HMI tags "Default tag table"
   "10_DI_DATA_5T1_PWR_OK" : Bool = PLC "10_DI_DATA".5T1_PWR_OK, 1 s
   "10_DI_DATA_6Q6_PWR_OK" : Bool = PLC "10_DI_DATA".6Q6_PWR_OK, 1 s
   "10_DI_DATA_CV341_CLSD" : Bool = PLC "10_DI_DATA".CV341_CLSD, 1 s
   "10_DI_DATA_CV341_OPN" : Bool = PLC "10_DI_DATA".CV341_OPN, 1 s
   "10_DI_DATA_CV358_CLSD" : Bool = PLC "10_DI_DATA".CV358_CLSD, 1 s
   "10_DI_DATA_CV358_OPN" : Bool = PLC "10_DI_DATA".CV358_OPN, 1 s
   "10_DI_DATA_CV406_CLSD" : Bool = PLC "10_DI_DATA".CV406_CLSD, 1 s
   "10_DI_DATA_CV406_OPN" : Bool = PLC "10_DI_DATA".CV406_OPN, 1 s
   "10_DI_DATA_CV407_CLSD" : Bool = PLC "10_DI_DATA".CV407_CLSD, 1 s
   "10_DI_DATA_CV407_OPN" : Bool = PLC "10_DI_DATA".CV407_OPN, 1 s
   "10_DI_DATA_CV409_CLSD" : Bool = PLC "10_DI_DATA".CV409_CLSD, 1 s
   "10_DI_DATA_CV409_OPN" : Bool = PLC "10_DI_DATA".CV409_OPN, 1 s
   "10_DI_DATA_CV411_CLSD" : Bool = PLC "10_DI_DATA".CV411_CLSD, 1 s
   "10_DI_DATA_CV411_OPN" : Bool = PLC "10_DI_DATA".CV411_OPN, 1 s
   "10_DI_DATA_CV441_CLSD" : Bool = PLC "10_DI_DATA".CV441_CLSD, 1 s
   "10_DI_DATA_CV441_OPN" : Bool = PLC "10_DI_DATA".CV441_OPN, 1 s
   "10_DI_DATA_E_400_NOK" : Bool = PLC "10_DI_DATA".E_400_NOK, 1 s
   "10_DI_DATA_E_400_RUN" : Bool = PLC "10_DI_DATA".E_400_RUN, 1 s
   "10_DI_DATA_E_400_SHTDN" : Bool = PLC "10_DI_DATA".E_400_SHTDN, 1 s
   "10_DI_DATA_E_400_STPD" : Bool = PLC "10_DI_DATA".E_400_STPD, 1 s
   "10_DI_DATA_EPB_8S1" : Bool = PLC "10_DI_DATA".EPB_8S1, 1 s
   "10_DI_DATA_FS_332 FLW_OK" : Bool = PLC "10_DI_DATA"."FS_332 FLW_OK", 1 s
   "10_DI_DATA_FS_350_FLW_OK" : Bool = PLC "10_DI_DATA".FS_350_FLW_OK, 1 s
   "10_DI_DATA_LS_303_LO" : Bool = PLC "10_DI_DATA".LS_303_LO, 1 s
   "10_DI_DATA_P_303_ENBLD" : Bool = PLC "10_DI_DATA".P_303_ENBLD, 1 s
   "10_DI_DATA_P_303_OK" : Bool = PLC "10_DI_DATA".P_303_OK, 1 s
   "10_DI_DATA_P_304_ENBLD" : Bool = PLC "10_DI_DATA".P_304_ENBLD, 1 s
   "10_DI_DATA_P_304_OK" : Bool = PLC "10_DI_DATA".P_304_OK, 1 s
   "10_DI_DATA_PB_10S1" : Bool = PLC "10_DI_DATA".PB_10S1, 1 s
   "10_DI_DATA_PB_10S2" : Bool = PLC "10_DI_DATA".PB_10S2, 1 s
   "10_DI_DATA_R3_SPR_DI_136_0" : Bool = PLC "10_DI_DATA".R3_SPR_DI_136_0, 1 s
   "10_DI_DATA_R3_SPR_DI_136_1" : Bool = PLC "10_DI_DATA".R3_SPR_DI_136_1, 1 s
   "100_BC_AUTO_SEQ_DB_CRNT_STEP" : Int = PLC "100_BC_AUTO_SEQ_DB".CRNT_STEP, 1 s
   "100_GCU_AUTO_SEQ_DB_CRNT_STEP" : Int = PLC "100_GCU_AUTO_SEQ_DB".CRNT_STEP, 1 s
   "100_GCU_AUTO_SEQ_DB_RNG" : Bool = PLC "100_GCU_AUTO_SEQ_DB".RNG, 1 s
   "100_IGG_AUTO_SEQ_DB_CRNT_STEP" : Int = PLC "100_IGG_AUTO_SEQ_DB".CRNT_STEP, 1 s
   "101_Fuel_Pumps_DB_Duty Is A" : Bool = PLC "101_Fuel_Pumps_DB"."Duty Is A", 1 s
   "101_Fuel_Pumps_DB_Duty Is B" : Bool = PLC "101_Fuel_Pumps_DB"."Duty Is B", 1 s
   "102_Pilot_Burner_DB_RUNNING" : Bool = PLC "102_Pilot_Burner_DB".RUNNING, 1 s
   "103_Main_Burner_DB_Days burn_CV" : Int = PLC "103_Main_Burner_DB"."Days burn".CV, 1 s
   "103_Main_Burner_DB_DN_OK" : Bool = PLC "103_Main_Burner_DB".DN_OK, 1 s
   "103_Main_Burner_DB_Hours burn_CV" : Int = PLC "103_Main_Burner_DB"."Hours burn".CV, 1 s
   "103_Main_Burner_DB_Minutes burn_CV" : Int = PLC "103_Main_Burner_DB"."Minutes burn".CV, 1 s
   "103_Main_Burner_DB_RUN" : Bool = PLC "103_Main_Burner_DB".RUN, 1 s
   "103_Main_Burner_DB_RUNNING" : Bool = PLC "103_Main_Burner_DB".RUNNING, 1 s
   "103_Main_Burner_DB_Seconds burn_CV" : Int = PLC "103_Main_Burner_DB"."Seconds burn".CV, 1 s
   "103_Main_Burner_DB_STATE" : Int = PLC "103_Main_Burner_DB".STATE, 1 s
   "103_Main_Burner_DB_Status" : Int = PLC "103_Main_Burner_DB".Status, 1 s
   "1111_PID_CV111_Setpoint" : Real = PLC "1111_PID_CV111".Setpoint, 1 s
   "12_AI_Data_CV_405_SCALED" : Real = PLC "12_AI_Data".CV_405_SCALED, 1 s
   "12_AI_Data_E_400_PT002_SCALED" : Real = PLC "12_AI_Data".E_400_PT002_SCALED, 1 s
   "12_AI_Data_E_400_TE002_SCALED" : Real = PLC "12_AI_Data".E_400_TE002_SCALED, 1 s
   "12_AI_Data_LIT_304_SCALED" : Real = PLC "12_AI_Data".LIT_304_SCALED, 1 s
   "12_AI_Data_PIT_348_SCALED" : Real = PLC "12_AI_Data".PIT_348_SCALED, 1 s
   "12_AI_Data_PIT_353_SCALED" : Real = PLC "12_AI_Data".PIT_353_SCALED, 1 s
   "12_AI_Data_PIT_358_SCALED" : Real = PLC "12_AI_Data".PIT_358_SCALED, 1 s
   "12_AI_Data_PIT_416_SCALED" : Real = PLC "12_AI_Data".PIT_416_SCALED, 1 s
   "12_AI_Data_R3_SPR_AI_802_SCALED" : Real = PLC "12_AI_Data".R3_SPR_AI_802_SCALED, 1 s
   "12_AI_Data_R3_SPR_AI_824_SCALED" : Real = PLC "12_AI_Data".R3_SPR_AI_824_SCALED, 1 s
   "12_AI_Data_R3_SPR_AI_826_SCALED" : Real = PLC "12_AI_Data".R3_SPR_AI_826_SCALED, 1 s
   "12_AI_Data_R3_SPR_AI_828_SCALED" : Real = PLC "12_AI_Data".R3_SPR_AI_828_SCALED, 1 s
   "12_AI_Data_R3_SPR_AI_830_SCALED" : Real = PLC "12_AI_Data".R3_SPR_AI_830_SCALED, 1 s
   "12_AI_Data_SL_400_SCALED" : Real = PLC "12_AI_Data".SL_400_SCALED, 1 s
   "12_AI_Data_TIT_406_SCALED" : Real = PLC "12_AI_Data".TIT_406_SCALED, 1 s
   "12_AI_Data_TIT_408_SCALED" : Real = PLC "12_AI_Data".TIT_408_SCALED, 1 s
   "14_DQ_DATA_13P1" : Bool = PLC "14_DQ_DATA".13P1, 1 s
   "14_DQ_DATA_13P2" : Bool = PLC "14_DQ_DATA".13P2, 1 s
   "14_DQ_DATA_13P3" : Bool = PLC "14_DQ_DATA".13P3, 1 s
   "14_DQ_DATA_13P4" : Bool = PLC "14_DQ_DATA".13P4, 1 s
   "14_DQ_DATA_13P5" : Bool = PLC "14_DQ_DATA".13P5, 1 s
   "14_DQ_DATA_E_400_STP" : Bool = PLC "14_DQ_DATA".E_400_STP, 1 s
   "14_DQ_DATA_P_303" : Bool = PLC "14_DQ_DATA".P_303, 1 s
   "14_DQ_DATA_P_304" : Bool = PLC "14_DQ_DATA".P_304, 1 s
   "14_DQ_DATA_R3_SPR_DQ_138_7" : Bool = PLC "14_DQ_DATA".R3_SPR_DQ_138_7, 1 s
   "14_DQ_DATA_R3_SPR_DQ_139_7" : Bool = PLC "14_DQ_DATA".R3_SPR_DQ_139_7, 1 s
   "140_PGC_HRS_RUN_DB_HRS" : Int = PLC "140_PGC_HRS_RUN_DB".HRS, 1 s
   "140_PGC_HRS_RUN_DB_MINS" : Int = PLC "140_PGC_HRS_RUN_DB".MINS, 1 s
   "140_PGC_HRS_RUN_DB_RST" : Bool = PLC "140_PGC_HRS_RUN_DB".RST, 1 s
   "140_PGC_HRS_RUN_DB_SECS" : Int = PLC "140_PGC_HRS_RUN_DB".SECS, 1 s
   "140_PGC_HRS_RUN_DB_SHRS_IP" : Int = PLC "140_PGC_HRS_RUN_DB".SHRS_IP, 1 s
   "140_PGC_HRS_RUN_DB_SRV_HRS" : Int = PLC "140_PGC_HRS_RUN_DB".SRV_HRS, 1 s
   "140_PGC_HRS_RUN_DB_SRVC" : Bool = PLC "140_PGC_HRS_RUN_DB".SRVC, 1 s
   "1405_PID_CV405_CtrlParamsBackUp_Gain" : Real = PLC "1405_PID_CV405".CtrlParamsBackUp.Gain, 1 s
   "1405_PID_CV405_CtrlParamsBackUp_Ti" : Real = PLC "1405_PID_CV405".CtrlParamsBackUp.Ti, 1 s
   "150_GCU_LCL_CNTRL_DB_LCL_CNTRL_ACTV" : Bool = PLC "150_GCU_LCL_CNTRL_DB".LCL_CNTRL_ACTV, 1 s
   "150_GCU_LCL_CNTRL_DB_OPN_ACTV_GTT_VLVS" : Bool = PLC "150_GCU_LCL_CNTRL_DB".OPN_ACTV_GTT_VLVS, 1 s
   "150_GCU_LCL_CNTRL_DB_RUN_WITH_AIR" : Bool = PLC "150_GCU_LCL_CNTRL_DB".RUN_WITH_AIR, 1 s
   "150_GCU_LCL_CNTRL_DB_RUN_WITH_IG" : Bool = PLC "150_GCU_LCL_CNTRL_DB".RUN_WITH_IG, 1 s
   "150_GCU_LCL_CNTRL_DB_STOP" : Bool = PLC "150_GCU_LCL_CNTRL_DB".STOP, 1 s
   "150_GCU_LCL_CNTRL_DB_STRT_AIR" : Bool = PLC "150_GCU_LCL_CNTRL_DB".STRT_AIR, 1 s
   "150_GCU_LCL_CNTRL_DB_STRT_IG" : Bool = PLC "150_GCU_LCL_CNTRL_DB".STRT_IG, 1 s
   "150_GCU_LCL_CNTRL_DB_SYS_OK_FOR_LCL" : Bool = PLC "150_GCU_LCL_CNTRL_DB".SYS_OK_FOR_LCL, 1 s
   "16_AQ_Data_CV405_CNTRL" : Real = PLC "16_AQ_Data".CV405_CNTRL, 1 s
   "19_AUTO_CMNDS_Data_CV203_RAMP_CNTRL" : Bool = PLC "19_AUTO_CMNDS_Data".CV203_RAMP_CNTRL, 1 s
   "19_AUTO_CMNDS_Data_CV405_PID_MDLTG" : Bool = PLC "19_AUTO_CMNDS_Data".CV405_PID_MDLTG, 1 s
   "19_AUTO_CMNDS_Data_LIT304_CMND_High" : Real = PLC "19_AUTO_CMNDS_Data".LIT304_CMND_High, 1 s
   "19_AUTO_CMNDS_Data_LIT304_CMND_HighHigh" : Real = PLC "19_AUTO_CMNDS_Data".LIT304_CMND_HighHigh, 1 s
   "19_AUTO_CMNDS_Data_LIT304_CMND_Low" : Real = PLC "19_AUTO_CMNDS_Data".LIT304_CMND_Low, 1 s
   "19_AUTO_CMNDS_Data_LIT304_CMND_LowLow" : Real = PLC "19_AUTO_CMNDS_Data".LIT304_CMND_LowLow, 1 s
   "19_AUTO_CMNDS_Data_LIT304_CMND_Target" : Real = PLC "19_AUTO_CMNDS_Data".LIT304_CMND_Target, 1 s
   "19_AUTO_CMNDS_Data_PIT353_CMND_High" : Real = PLC "19_AUTO_CMNDS_Data".PIT353_CMND_High, 1 s
   "19_AUTO_CMNDS_Data_PIT353_CMND_HighHigh" : Real = PLC "19_AUTO_CMNDS_Data".PIT353_CMND_HighHigh, 1 s
   "19_AUTO_CMNDS_Data_PIT353_CMND_Low" : Real = PLC "19_AUTO_CMNDS_Data".PIT353_CMND_Low, 1 s
   "19_AUTO_CMNDS_Data_PIT353_CMND_LowLow" : Real = PLC "19_AUTO_CMNDS_Data".PIT353_CMND_LowLow, 1 s
   "19_AUTO_CMNDS_Data_PIT358_CMND_High" : Real = PLC "19_AUTO_CMNDS_Data".PIT358_CMND_High, 1 s
   "19_AUTO_CMNDS_Data_PIT358_CMND_HighHigh" : Real = PLC "19_AUTO_CMNDS_Data".PIT358_CMND_HighHigh, 1 s
   "19_AUTO_CMNDS_Data_PIT358_CMND_Low" : Real = PLC "19_AUTO_CMNDS_Data".PIT358_CMND_Low, 1 s
   "19_AUTO_CMNDS_Data_PIT358_CMND_LowLow" : Real = PLC "19_AUTO_CMNDS_Data".PIT358_CMND_LowLow, 1 s
   "19_AUTO_CMNDS_Data_PIT416_CMND_Target" : Real = PLC "19_AUTO_CMNDS_Data".PIT416_CMND_Target, 1 s
   "20_TANKS_IP_DATA_RIO_01_FIRST_TANK_BWT_DO" : Real = PLC "20_TANKS_IP_DATA".RIO_01.FIRST_TANK.BWT_DO, 1 s
   "20_TANKS_IP_DATA_RIO_01_FIRST_TANK_BWT_LEVEL" : Real = PLC "20_TANKS_IP_DATA".RIO_01.FIRST_TANK.BWT_LEVEL, 1 s
   "20_TANKS_IP_DATA_RIO_01_FIRST_TANK_BWT_LEVEL_HIHI" : Bool = PLC "20_TANKS_IP_DATA".RIO_01.FIRST_TANK.BWT_LEVEL_HIHI, 1 s
   "20_TANKS_IP_DATA_RIO_01_FIRST_TANK_BWT_PH" : Real = PLC "20_TANKS_IP_DATA".RIO_01.FIRST_TANK.BWT_PH, 1 s
   "20_TANKS_IP_DATA_RIO_01_FIRST_TANK_BWT_TEMP" : Real = PLC "20_TANKS_IP_DATA".RIO_01.FIRST_TANK.BWT_TEMP, 1 s
   "20_TANKS_IP_DATA_RIO_01_FIRST_TANK_DECK_IG_PRESS" : Real = PLC "20_TANKS_IP_DATA".RIO_01.FIRST_TANK.DECK_IG_PRESS, 1 s
   "20_TANKS_IP_DATA_RIO_01_FIRST_TANK_GTT_ISOL_VALVE_CLSD" : Bool = PLC "20_TANKS_IP_DATA".RIO_01.FIRST_TANK.GTT_ISOL_VALVE_CLSD, 1 s
   "20_TANKS_IP_DATA_RIO_01_FIRST_TANK_GTT_ISOL_VALVE_OPEN" : Bool = PLC "20_TANKS_IP_DATA".RIO_01.FIRST_TANK.GTT_ISOL_VALVE_OPEN, 1 s
   "20_TANKS_IP_DATA_RIO_01_FIRST_TANK_MBG_FLOW" : Real = PLC "20_TANKS_IP_DATA".RIO_01.FIRST_TANK.MBG_FLOW, 1 s
   "20_TANKS_IP_DATA_RIO_01_FIRST_TANK_O2_MONITOR" : Real = PLC "20_TANKS_IP_DATA".RIO_01.FIRST_TANK.O2_MONITOR, 1 s
   "20_TANKS_IP_DATA_RIO_01_FIRST_TANK_TANKS_PRESS" : Real = PLC "20_TANKS_IP_DATA".RIO_01.FIRST_TANK.TANKS_PRESS, 1 s
   "20_TANKS_IP_DATA_RIO_01_FIRST_TANK_USD_FLOW" : Real = PLC "20_TANKS_IP_DATA".RIO_01.FIRST_TANK.USD_FLOW, 1 s
   "20_TANKS_IP_DATA_RIO_01_SECOND_TANK_BWT_DO" : Real = PLC "20_TANKS_IP_DATA".RIO_01.SECOND_TANK.BWT_DO, 1 s
   "20_TANKS_IP_DATA_RIO_01_SECOND_TANK_BWT_LEVEL" : Real = PLC "20_TANKS_IP_DATA".RIO_01.SECOND_TANK.BWT_LEVEL, 1 s
   "20_TANKS_IP_DATA_RIO_01_SECOND_TANK_BWT_LEVEL_HIHI" : Bool = PLC "20_TANKS_IP_DATA".RIO_01.SECOND_TANK.BWT_LEVEL_HIHI, 1 s
   "20_TANKS_IP_DATA_RIO_01_SECOND_TANK_BWT_PH" : Real = PLC "20_TANKS_IP_DATA".RIO_01.SECOND_TANK.BWT_PH, 1 s
   "20_TANKS_IP_DATA_RIO_01_SECOND_TANK_BWT_TEMP" : Real = PLC "20_TANKS_IP_DATA".RIO_01.SECOND_TANK.BWT_TEMP, 1 s
   "20_TANKS_IP_DATA_RIO_01_SECOND_TANK_GTT_ISOL_VALVE_CLSD" : Bool = PLC "20_TANKS_IP_DATA".RIO_01.SECOND_TANK.GTT_ISOL_VALVE_CLSD, 1 s
   "20_TANKS_IP_DATA_RIO_01_SECOND_TANK_GTT_ISOL_VALVE_OPEN" : Bool = PLC "20_TANKS_IP_DATA".RIO_01.SECOND_TANK.GTT_ISOL_VALVE_OPEN, 1 s
   "20_TANKS_IP_DATA_RIO_01_SECOND_TANK_MBG_FLOW" : Real = PLC "20_TANKS_IP_DATA".RIO_01.SECOND_TANK.MBG_FLOW, 1 s
   "20_TANKS_IP_DATA_RIO_01_SECOND_TANK_TANKS_PRESS" : Real = PLC "20_TANKS_IP_DATA".RIO_01.SECOND_TANK.TANKS_PRESS, 1 s
   "20_TANKS_IP_DATA_RIO_01_SECOND_TANK_USD_FLOW" : Real = PLC "20_TANKS_IP_DATA".RIO_01.SECOND_TANK.USD_FLOW, 1 s
   "20_TANKS_IP_DATA_RIO_01_THIRD_TANK_BWT_DO" : Real = PLC "20_TANKS_IP_DATA".RIO_01.THIRD_TANK.BWT_DO, 1 s
   "20_TANKS_IP_DATA_RIO_01_THIRD_TANK_BWT_LEVEL" : Real = PLC "20_TANKS_IP_DATA".RIO_01.THIRD_TANK.BWT_LEVEL, 1 s
   "20_TANKS_IP_DATA_RIO_01_THIRD_TANK_BWT_LEVEL_HIHI" : Bool = PLC "20_TANKS_IP_DATA".RIO_01.THIRD_TANK.BWT_LEVEL_HIHI, 1 s
   "20_TANKS_IP_DATA_RIO_01_THIRD_TANK_BWT_PH" : Real = PLC "20_TANKS_IP_DATA".RIO_01.THIRD_TANK.BWT_PH, 1 s
   "20_TANKS_IP_DATA_RIO_01_THIRD_TANK_BWT_TEMP" : Real = PLC "20_TANKS_IP_DATA".RIO_01.THIRD_TANK.BWT_TEMP, 1 s
   "20_TANKS_IP_DATA_RIO_01_THIRD_TANK_DECK_IG_PRESS" : Real = PLC "20_TANKS_IP_DATA".RIO_01.THIRD_TANK.DECK_IG_PRESS, 1 s
   "20_TANKS_IP_DATA_RIO_01_THIRD_TANK_GTT_ISOL_VALVE_CLSD" : Bool = PLC "20_TANKS_IP_DATA".RIO_01.THIRD_TANK.GTT_ISOL_VALVE_CLSD, 1 s
   "20_TANKS_IP_DATA_RIO_01_THIRD_TANK_GTT_ISOL_VALVE_OPEN" : Bool = PLC "20_TANKS_IP_DATA".RIO_01.THIRD_TANK.GTT_ISOL_VALVE_OPEN, 1 s
   "20_TANKS_IP_DATA_RIO_01_THIRD_TANK_MBG_FLOW" : Real = PLC "20_TANKS_IP_DATA".RIO_01.THIRD_TANK.MBG_FLOW, 1 s
   "20_TANKS_IP_DATA_RIO_01_THIRD_TANK_O2_MONITOR" : Real = PLC "20_TANKS_IP_DATA".RIO_01.THIRD_TANK.O2_MONITOR, 1 s
   "20_TANKS_IP_DATA_RIO_01_THIRD_TANK_TANKS_PRESS" : Real = PLC "20_TANKS_IP_DATA".RIO_01.THIRD_TANK.TANKS_PRESS, 1 s
   "20_TANKS_IP_DATA_RIO_01_THIRD_TANK_USD_FLOW" : Real = PLC "20_TANKS_IP_DATA".RIO_01.THIRD_TANK.USD_FLOW, 1 s
   "20_TANKS_IP_DATA_RIO_02_FIRST_TANK_BWT_DO" : Real = PLC "20_TANKS_IP_DATA".RIO_02.FIRST_TANK.BWT_DO, 1 s
   "20_TANKS_IP_DATA_RIO_02_FIRST_TANK_BWT_LEVEL" : Real = PLC "20_TANKS_IP_DATA".RIO_02.FIRST_TANK.BWT_LEVEL, 1 s
   "20_TANKS_IP_DATA_RIO_02_FIRST_TANK_BWT_LEVEL_HIHI" : Bool = PLC "20_TANKS_IP_DATA".RIO_02.FIRST_TANK.BWT_LEVEL_HIHI AT %DB1.DBW0, 1 s
   "20_TANKS_IP_DATA_RIO_02_FIRST_TANK_BWT_PH" : Real = PLC "20_TANKS_IP_DATA".RIO_02.FIRST_TANK.BWT_PH, 1 s
   "20_TANKS_IP_DATA_RIO_02_FIRST_TANK_BWT_TEMP" : Real = PLC "20_TANKS_IP_DATA".RIO_02.FIRST_TANK.BWT_TEMP, 1 s
   "20_TANKS_IP_DATA_RIO_02_FIRST_TANK_DECK_IG_PRESS" : Real = PLC "20_TANKS_IP_DATA".RIO_02.FIRST_TANK.DECK_IG_PRESS, 1 s
   "20_TANKS_IP_DATA_RIO_02_FIRST_TANK_GTT_ISOL_VALVE_CLSD" : Bool = PLC "20_TANKS_IP_DATA".RIO_02.FIRST_TANK.GTT_ISOL_VALVE_CLSD AT %DB1.DBW0, 1 s
   "20_TANKS_IP_DATA_RIO_02_FIRST_TANK_GTT_ISOL_VALVE_OPEN" : Bool = PLC "20_TANKS_IP_DATA".RIO_02.FIRST_TANK.GTT_ISOL_VALVE_OPEN AT %DB1.DBW0, 1 s
   "20_TANKS_IP_DATA_RIO_02_FIRST_TANK_MBG_FLOW" : Real = PLC "20_TANKS_IP_DATA".RIO_02.FIRST_TANK.MBG_FLOW AT %DB1.DBW0, 1 s
   "20_TANKS_IP_DATA_RIO_02_FIRST_TANK_MBG_FLOW_raw" : Real = PLC "20_TANKS_IP_DATA".RIO_02.FIRST_TANK."MBG_FLOW N" AT %DB1.DBD0, 1 s
   "20_TANKS_IP_DATA_RIO_02_FIRST_TANK_O2_MONITOR" : Real = PLC "20_TANKS_IP_DATA".RIO_02.FIRST_TANK.O2_MONITOR AT %DB1.DBW0, 1 s
   "20_TANKS_IP_DATA_RIO_02_FIRST_TANK_TANK_VENT_A_CLSD" : Bool = PLC "20_TANKS_IP_DATA".RIO_02.FIRST_TANK.TANK_VENT_A_CLSD AT %DB1.DBW0, 1 s
   "20_TANKS_IP_DATA_RIO_02_FIRST_TANK_TANK_VENT_A_OPEN" : Bool = PLC "20_TANKS_IP_DATA".RIO_02.FIRST_TANK.TANK_VENT_A_OPEN AT %DB1.DBW0, 1 s
   "20_TANKS_IP_DATA_RIO_02_FIRST_TANK_TANK_VENT_B_CLSD" : Bool = PLC "20_TANKS_IP_DATA".RIO_02.FIRST_TANK.TANK_VENT_B_CLSD AT %DB1.DBW0, 1 s
   "20_TANKS_IP_DATA_RIO_02_FIRST_TANK_TANK_VENT_B_OPEN" : Bool = PLC "20_TANKS_IP_DATA".RIO_02.FIRST_TANK.TANK_VENT_B_OPEN AT %DB1.DBW0, 1 s
   "20_TANKS_IP_DATA_RIO_02_FIRST_TANK_TANKS_PRESS" : Real = PLC "20_TANKS_IP_DATA".RIO_02.FIRST_TANK.TANKS_PRESS AT %DB1.DBW0, 1 s
   "20_TANKS_IP_DATA_RIO_02_FIRST_TANK_TANKS_PRESS_HIHI" : Bool = PLC "20_TANKS_IP_DATA".RIO_02.FIRST_TANK.TANKS_PRESS_HIHI AT %DB1.DBW0, 1 s
   "20_TANKS_IP_DATA_RIO_02_FIRST_TANK_USD_FLOW" : Real = PLC "20_TANKS_IP_DATA".RIO_02.FIRST_TANK.USD_FLOW AT %DB1.DBW0, 1 s
   "20_TANKS_IP_DATA_RIO_02_FIRST_TANK_USD_FLOW_raw" : Real = PLC "20_TANKS_IP_DATA".RIO_02.FIRST_TANK."USD FLOW  N" AT %DB1.DBD0, 1 s
   "20_TANKS_IP_DATA_RIO_02_SECOND_TANK_BWT_DO" : Real = PLC "20_TANKS_IP_DATA".RIO_02.SECOND_TANK.BWT_DO, 1 s
   "20_TANKS_IP_DATA_RIO_02_SECOND_TANK_BWT_LEVEL" : Real = PLC "20_TANKS_IP_DATA".RIO_02.SECOND_TANK.BWT_LEVEL, 1 s
   "20_TANKS_IP_DATA_RIO_02_SECOND_TANK_BWT_LEVEL_HIHI" : Bool = PLC "20_TANKS_IP_DATA".RIO_02.SECOND_TANK.BWT_LEVEL_HIHI AT %DB1.DBW0, 1 s
   "20_TANKS_IP_DATA_RIO_02_SECOND_TANK_BWT_PH" : Real = PLC "20_TANKS_IP_DATA".RIO_02.SECOND_TANK.BWT_PH, 1 s
   "20_TANKS_IP_DATA_RIO_02_SECOND_TANK_BWT_TEMP" : Real = PLC "20_TANKS_IP_DATA".RIO_02.SECOND_TANK.BWT_TEMP, 1 s
   "20_TANKS_IP_DATA_RIO_02_SECOND_TANK_DECK_IG_PRESS" : Real = PLC "20_TANKS_IP_DATA".RIO_02.SECOND_TANK.DECK_IG_PRESS AT %DB1.DBW0, 1 s
   "20_TANKS_IP_DATA_RIO_02_SECOND_TANK_GTT_ISOL_VALVE_CLSD" : Bool = PLC "20_TANKS_IP_DATA".RIO_02.SECOND_TANK.GTT_ISOL_VALVE_CLSD AT %DB1.DBW0, 1 s
   "20_TANKS_IP_DATA_RIO_02_SECOND_TANK_GTT_ISOL_VALVE_OPEN" : Bool = PLC "20_TANKS_IP_DATA".RIO_02.SECOND_TANK.GTT_ISOL_VALVE_OPEN AT %DB1.DBW0, 1 s
   "20_TANKS_IP_DATA_RIO_02_SECOND_TANK_MBG_FLOW" : Real = PLC "20_TANKS_IP_DATA".RIO_02.SECOND_TANK.MBG_FLOW AT %DB1.DBW0, 1 s
   "20_TANKS_IP_DATA_RIO_02_SECOND_TANK_MBG_FLOW_raw" : Real = PLC "20_TANKS_IP_DATA".RIO_02.SECOND_TANK."MBG_FLOW N" AT %DB1.DBD0, 1 s
   "20_TANKS_IP_DATA_RIO_02_SECOND_TANK_O2_MONITOR" : Real = PLC "20_TANKS_IP_DATA".RIO_02.SECOND_TANK.O2_MONITOR AT %DB1.DBW0, 1 s
   "20_TANKS_IP_DATA_RIO_02_SECOND_TANK_TANK_VENT_A_CLSD" : Bool = PLC "20_TANKS_IP_DATA".RIO_02.SECOND_TANK.TANK_VENT_A_CLSD AT %DB1.DBW0, 1 s
   "20_TANKS_IP_DATA_RIO_02_SECOND_TANK_TANK_VENT_A_OPEN" : Bool = PLC "20_TANKS_IP_DATA".RIO_02.SECOND_TANK.TANK_VENT_A_OPEN AT %DB1.DBW0, 1 s
   "20_TANKS_IP_DATA_RIO_02_SECOND_TANK_TANK_VENT_B_CLSD" : Bool = PLC "20_TANKS_IP_DATA".RIO_02.SECOND_TANK.TANK_VENT_B_CLSD AT %DB1.DBW0, 1 s
   "20_TANKS_IP_DATA_RIO_02_SECOND_TANK_TANK_VENT_B_OPEN" : Bool = PLC "20_TANKS_IP_DATA".RIO_02.SECOND_TANK.TANK_VENT_B_OPEN AT %DB1.DBW0, 1 s
   "20_TANKS_IP_DATA_RIO_02_SECOND_TANK_TANKS_PRESS" : Real = PLC "20_TANKS_IP_DATA".RIO_02.SECOND_TANK.TANKS_PRESS AT %DB1.DBW0, 1 s
   "20_TANKS_IP_DATA_RIO_02_SECOND_TANK_TANKS_PRESS_HIHI" : Bool = PLC "20_TANKS_IP_DATA".RIO_02.SECOND_TANK.TANKS_PRESS_HIHI AT %DB1.DBW0, 1 s
   "20_TANKS_IP_DATA_RIO_02_SECOND_TANK_USD_FLOW" : Real = PLC "20_TANKS_IP_DATA".RIO_02.SECOND_TANK.USD_FLOW AT %DB1.DBW0, 1 s
   "20_TANKS_IP_DATA_RIO_02_SECOND_TANK_USD_FLOW_raw" : Real = PLC "20_TANKS_IP_DATA".RIO_02.SECOND_TANK."USD FLOW  N" AT %DB1.DBD0, 1 s
   "20_TANKS_IP_DATA_RIO_03_FIRST_TANK_BWT_DO" : Real = PLC "20_TANKS_IP_DATA".RIO_03.FIRST_TANK.BWT_DO, 1 s
   "20_TANKS_IP_DATA_RIO_03_FIRST_TANK_BWT_LEVEL" : Real = PLC "20_TANKS_IP_DATA".RIO_03.FIRST_TANK.BWT_LEVEL, 1 s
   "20_TANKS_IP_DATA_RIO_03_FIRST_TANK_BWT_LEVEL_HIHI" : Bool = PLC "20_TANKS_IP_DATA".RIO_03.FIRST_TANK.BWT_LEVEL_HIHI, 1 s
   "20_TANKS_IP_DATA_RIO_03_FIRST_TANK_BWT_PH" : Real = PLC "20_TANKS_IP_DATA".RIO_03.FIRST_TANK.BWT_PH, 1 s
   "20_TANKS_IP_DATA_RIO_03_FIRST_TANK_BWT_TEMP" : Real = PLC "20_TANKS_IP_DATA".RIO_03.FIRST_TANK.BWT_TEMP, 1 s
   "20_TANKS_IP_DATA_RIO_03_FIRST_TANK_DECK_IG_PRESS" : Real = PLC "20_TANKS_IP_DATA".RIO_03.FIRST_TANK.DECK_IG_PRESS, 1 s
   "20_TANKS_IP_DATA_RIO_03_FIRST_TANK_GTT_ISOL_VALVE_CLSD" : Bool = PLC "20_TANKS_IP_DATA".RIO_03.FIRST_TANK.GTT_ISOL_VALVE_CLSD, 1 s
   "20_TANKS_IP_DATA_RIO_03_FIRST_TANK_GTT_ISOL_VALVE_OPEN" : Bool = PLC "20_TANKS_IP_DATA".RIO_03.FIRST_TANK.GTT_ISOL_VALVE_OPEN, 1 s
   "20_TANKS_IP_DATA_RIO_03_FIRST_TANK_MBG_FLOW" : Real = PLC "20_TANKS_IP_DATA".RIO_03.FIRST_TANK.MBG_FLOW, 1 s
   "20_TANKS_IP_DATA_RIO_03_FIRST_TANK_O2_MONITOR" : Real = PLC "20_TANKS_IP_DATA".RIO_03.FIRST_TANK.O2_MONITOR, 1 s
   "20_TANKS_IP_DATA_RIO_03_FIRST_TANK_TANKS_PRESS" : Real = PLC "20_TANKS_IP_DATA".RIO_03.FIRST_TANK.TANKS_PRESS, 1 s
   "20_TANKS_IP_DATA_RIO_03_FIRST_TANK_USD_FLOW" : Real = PLC "20_TANKS_IP_DATA".RIO_03.FIRST_TANK.USD_FLOW, 1 s
   "20_TANKS_IP_DATA_RIO_03_SECOND_TANK_BWT_DO" : Real = PLC "20_TANKS_IP_DATA".RIO_03.SECOND_TANK.BWT_DO, 1 s
   "20_TANKS_IP_DATA_RIO_03_SECOND_TANK_BWT_LEVEL" : Real = PLC "20_TANKS_IP_DATA".RIO_03.SECOND_TANK.BWT_LEVEL, 1 s
   "20_TANKS_IP_DATA_RIO_03_SECOND_TANK_BWT_LEVEL_HIHI" : Bool = PLC "20_TANKS_IP_DATA".RIO_03.SECOND_TANK.BWT_LEVEL_HIHI, 1 s
   "20_TANKS_IP_DATA_RIO_03_SECOND_TANK_BWT_PH" : Real = PLC "20_TANKS_IP_DATA".RIO_03.SECOND_TANK.BWT_PH, 1 s
   "20_TANKS_IP_DATA_RIO_03_SECOND_TANK_BWT_TEMP" : Real = PLC "20_TANKS_IP_DATA".RIO_03.SECOND_TANK.BWT_TEMP, 1 s
   "20_TANKS_IP_DATA_RIO_03_SECOND_TANK_GTT_ISOL_VALVE_CLSD" : Bool = PLC "20_TANKS_IP_DATA".RIO_03.SECOND_TANK.GTT_ISOL_VALVE_CLSD, 1 s
   "20_TANKS_IP_DATA_RIO_03_SECOND_TANK_GTT_ISOL_VALVE_OPEN" : Bool = PLC "20_TANKS_IP_DATA".RIO_03.SECOND_TANK.GTT_ISOL_VALVE_OPEN, 1 s
   "20_TANKS_IP_DATA_RIO_03_SECOND_TANK_MBG_FLOW" : Real = PLC "20_TANKS_IP_DATA".RIO_03.SECOND_TANK.MBG_FLOW, 1 s
   "20_TANKS_IP_DATA_RIO_03_SECOND_TANK_O2_MONITOR" : Real = PLC "20_TANKS_IP_DATA".RIO_03.SECOND_TANK.O2_MONITOR, 1 s
   "20_TANKS_IP_DATA_RIO_03_SECOND_TANK_TANKS_PRESS" : Real = PLC "20_TANKS_IP_DATA".RIO_03.SECOND_TANK.TANKS_PRESS, 1 s
   "20_TANKS_IP_DATA_RIO_03_SECOND_TANK_USD_FLOW" : Real = PLC "20_TANKS_IP_DATA".RIO_03.SECOND_TANK.USD_FLOW, 1 s
   "20_TANKS_IP_DATA_RIO_04_FIRST_TANK_BWT_DO" : Real = PLC "20_TANKS_IP_DATA".RIO_04.FIRST_TANK.BWT_DO, 1 s
   "20_TANKS_IP_DATA_RIO_04_FIRST_TANK_BWT_LEVEL" : Real = PLC "20_TANKS_IP_DATA".RIO_04.FIRST_TANK.BWT_LEVEL, 1 s
   "20_TANKS_IP_DATA_RIO_04_FIRST_TANK_BWT_LEVEL_HIHI" : Bool = PLC "20_TANKS_IP_DATA".RIO_04.FIRST_TANK.BWT_LEVEL_HIHI, 1 s
   "20_TANKS_IP_DATA_RIO_04_FIRST_TANK_BWT_PH" : Real = PLC "20_TANKS_IP_DATA".RIO_04.FIRST_TANK.BWT_PH, 1 s
   "20_TANKS_IP_DATA_RIO_04_FIRST_TANK_BWT_TEMP" : Real = PLC "20_TANKS_IP_DATA".RIO_04.FIRST_TANK.BWT_TEMP, 1 s
   "20_TANKS_IP_DATA_RIO_04_FIRST_TANK_DECK_IG_PRESS" : Real = PLC "20_TANKS_IP_DATA".RIO_04.FIRST_TANK.DECK_IG_PRESS, 1 s
   "20_TANKS_IP_DATA_RIO_04_FIRST_TANK_GTT_ISOL_VALVE_CLSD" : Bool = PLC "20_TANKS_IP_DATA".RIO_04.FIRST_TANK.GTT_ISOL_VALVE_CLSD, 1 s
   "20_TANKS_IP_DATA_RIO_04_FIRST_TANK_GTT_ISOL_VALVE_OPEN" : Bool = PLC "20_TANKS_IP_DATA".RIO_04.FIRST_TANK.GTT_ISOL_VALVE_OPEN, 1 s
   "20_TANKS_IP_DATA_RIO_04_FIRST_TANK_MBG_FLOW" : Real = PLC "20_TANKS_IP_DATA".RIO_04.FIRST_TANK.MBG_FLOW, 1 s
   "20_TANKS_IP_DATA_RIO_04_FIRST_TANK_O2_MONITOR" : Real = PLC "20_TANKS_IP_DATA".RIO_04.FIRST_TANK.O2_MONITOR, 1 s
   "20_TANKS_IP_DATA_RIO_04_FIRST_TANK_TANKS_PRESS" : Real = PLC "20_TANKS_IP_DATA".RIO_04.FIRST_TANK.TANKS_PRESS, 1 s
   "20_TANKS_IP_DATA_RIO_04_FIRST_TANK_USD_FLOW" : Real = PLC "20_TANKS_IP_DATA".RIO_04.FIRST_TANK.USD_FLOW, 1 s
   "20_TANKS_IP_DATA_RIO_04_SECOND_TANK_BWT_DO" : Real = PLC "20_TANKS_IP_DATA".RIO_04.SECOND_TANK.BWT_DO, 1 s
   "20_TANKS_IP_DATA_RIO_04_SECOND_TANK_BWT_LEVEL" : Real = PLC "20_TANKS_IP_DATA".RIO_04.SECOND_TANK.BWT_LEVEL, 1 s
   "20_TANKS_IP_DATA_RIO_04_SECOND_TANK_BWT_LEVEL_HIHI" : Bool = PLC "20_TANKS_IP_DATA".RIO_04.SECOND_TANK.BWT_LEVEL_HIHI, 1 s
   "20_TANKS_IP_DATA_RIO_04_SECOND_TANK_BWT_PH" : Real = PLC "20_TANKS_IP_DATA".RIO_04.SECOND_TANK.BWT_PH, 1 s
   "20_TANKS_IP_DATA_RIO_04_SECOND_TANK_BWT_TEMP" : Real = PLC "20_TANKS_IP_DATA".RIO_04.SECOND_TANK.BWT_TEMP, 1 s
   "20_TANKS_IP_DATA_RIO_04_SECOND_TANK_GTT_ISOL_VALVE_CLSD" : Bool = PLC "20_TANKS_IP_DATA".RIO_04.SECOND_TANK.GTT_ISOL_VALVE_CLSD, 1 s
   "20_TANKS_IP_DATA_RIO_04_SECOND_TANK_GTT_ISOL_VALVE_OPEN" : Bool = PLC "20_TANKS_IP_DATA".RIO_04.SECOND_TANK.GTT_ISOL_VALVE_OPEN, 1 s
   "20_TANKS_IP_DATA_RIO_04_SECOND_TANK_MBG_FLOW" : Real = PLC "20_TANKS_IP_DATA".RIO_04.SECOND_TANK.MBG_FLOW, 1 s
   "20_TANKS_IP_DATA_RIO_04_SECOND_TANK_O2_MONITOR" : Real = PLC "20_TANKS_IP_DATA".RIO_04.SECOND_TANK.O2_MONITOR, 1 s
   "20_TANKS_IP_DATA_RIO_04_SECOND_TANK_TANKS_PRESS" : Real = PLC "20_TANKS_IP_DATA".RIO_04.SECOND_TANK.TANKS_PRESS, 1 s
   "20_TANKS_IP_DATA_RIO_04_SECOND_TANK_USD_FLOW" : Real = PLC "20_TANKS_IP_DATA".RIO_04.SECOND_TANK.USD_FLOW, 1 s
   "20_TANKS_IP_DATA_RIO_05_FIRST_TANK_BWT_DO" : Real = PLC "20_TANKS_IP_DATA".RIO_05.FIRST_TANK.BWT_DO, 1 s
   "20_TANKS_IP_DATA_RIO_05_FIRST_TANK_BWT_LEVEL" : Real = PLC "20_TANKS_IP_DATA".RIO_05.FIRST_TANK.BWT_LEVEL, 1 s
   "20_TANKS_IP_DATA_RIO_05_FIRST_TANK_BWT_LEVEL_HIHI" : Bool = PLC "20_TANKS_IP_DATA".RIO_05.FIRST_TANK.BWT_LEVEL_HIHI, 1 s
   "20_TANKS_IP_DATA_RIO_05_FIRST_TANK_BWT_PH" : Real = PLC "20_TANKS_IP_DATA".RIO_05.FIRST_TANK.BWT_PH, 1 s
   "20_TANKS_IP_DATA_RIO_05_FIRST_TANK_BWT_TEMP" : Real = PLC "20_TANKS_IP_DATA".RIO_05.FIRST_TANK.BWT_TEMP, 1 s
   "20_TANKS_IP_DATA_RIO_05_FIRST_TANK_DECK_IG_PRESS" : Real = PLC "20_TANKS_IP_DATA".RIO_05.FIRST_TANK.DECK_IG_PRESS, 1 s
   "20_TANKS_IP_DATA_RIO_05_FIRST_TANK_GTT_ISOL_VALVE_CLSD" : Bool = PLC "20_TANKS_IP_DATA".RIO_05.FIRST_TANK.GTT_ISOL_VALVE_CLSD, 1 s
   "20_TANKS_IP_DATA_RIO_05_FIRST_TANK_GTT_ISOL_VALVE_OPEN" : Bool = PLC "20_TANKS_IP_DATA".RIO_05.FIRST_TANK.GTT_ISOL_VALVE_OPEN, 1 s
   "20_TANKS_IP_DATA_RIO_05_FIRST_TANK_MBG_FLOW" : Real = PLC "20_TANKS_IP_DATA".RIO_05.FIRST_TANK.MBG_FLOW, 1 s
   "20_TANKS_IP_DATA_RIO_05_FIRST_TANK_O2_MONITOR" : Real = PLC "20_TANKS_IP_DATA".RIO_05.FIRST_TANK.O2_MONITOR, 1 s
   "20_TANKS_IP_DATA_RIO_05_FIRST_TANK_TANKS_PRESS" : Real = PLC "20_TANKS_IP_DATA".RIO_05.FIRST_TANK.TANKS_PRESS, 1 s
   "20_TANKS_IP_DATA_RIO_05_FIRST_TANK_USD_FLOW" : Real = PLC "20_TANKS_IP_DATA".RIO_05.FIRST_TANK.USD_FLOW, 1 s
   "20_TANKS_IP_DATA_RIO_05_SECOND_TANK_BWT_DO" : Real = PLC "20_TANKS_IP_DATA".RIO_05.SECOND_TANK.BWT_DO, 1 s
   "20_TANKS_IP_DATA_RIO_05_SECOND_TANK_BWT_LEVEL" : Real = PLC "20_TANKS_IP_DATA".RIO_05.SECOND_TANK.BWT_LEVEL, 1 s
   "20_TANKS_IP_DATA_RIO_05_SECOND_TANK_BWT_LEVEL_HIHI" : Bool = PLC "20_TANKS_IP_DATA".RIO_05.SECOND_TANK.BWT_LEVEL_HIHI, 1 s
   "20_TANKS_IP_DATA_RIO_05_SECOND_TANK_BWT_PH" : Real = PLC "20_TANKS_IP_DATA".RIO_05.SECOND_TANK.BWT_PH, 1 s
   "20_TANKS_IP_DATA_RIO_05_SECOND_TANK_BWT_TEMP" : Real = PLC "20_TANKS_IP_DATA".RIO_05.SECOND_TANK.BWT_TEMP, 1 s
   "20_TANKS_IP_DATA_RIO_05_SECOND_TANK_GTT_ISOL_VALVE_CLSD" : Bool = PLC "20_TANKS_IP_DATA".RIO_05.SECOND_TANK.GTT_ISOL_VALVE_CLSD, 1 s
   "20_TANKS_IP_DATA_RIO_05_SECOND_TANK_GTT_ISOL_VALVE_OPEN" : Bool = PLC "20_TANKS_IP_DATA".RIO_05.SECOND_TANK.GTT_ISOL_VALVE_OPEN, 1 s
   "20_TANKS_IP_DATA_RIO_05_SECOND_TANK_MBG_FLOW" : Real = PLC "20_TANKS_IP_DATA".RIO_05.SECOND_TANK.MBG_FLOW, 1 s
   "20_TANKS_IP_DATA_RIO_05_SECOND_TANK_O2_MONITOR" : Real = PLC "20_TANKS_IP_DATA".RIO_05.SECOND_TANK.O2_MONITOR, 1 s
   "20_TANKS_IP_DATA_RIO_05_SECOND_TANK_TANKS_PRESS" : Real = PLC "20_TANKS_IP_DATA".RIO_05.SECOND_TANK.TANKS_PRESS, 1 s
   "20_TANKS_IP_DATA_RIO_05_SECOND_TANK_USD_FLOW" : Real = PLC "20_TANKS_IP_DATA".RIO_05.SECOND_TANK.USD_FLOW, 1 s
   "20_TANKS_IP_DATA_RIO_06_FIRST_TANK_BWT_DO" : Real = PLC "20_TANKS_IP_DATA".RIO_06.FIRST_TANK.BWT_DO, 1 s
   "20_TANKS_IP_DATA_RIO_06_FIRST_TANK_BWT_LEVEL" : Real = PLC "20_TANKS_IP_DATA".RIO_06.FIRST_TANK.BWT_LEVEL, 1 s
   "20_TANKS_IP_DATA_RIO_06_FIRST_TANK_BWT_LEVEL_HIHI" : Bool = PLC "20_TANKS_IP_DATA".RIO_06.FIRST_TANK.BWT_LEVEL_HIHI, 1 s
   "20_TANKS_IP_DATA_RIO_06_FIRST_TANK_BWT_PH" : Real = PLC "20_TANKS_IP_DATA".RIO_06.FIRST_TANK.BWT_PH, 1 s
   "20_TANKS_IP_DATA_RIO_06_FIRST_TANK_BWT_TEMP" : Real = PLC "20_TANKS_IP_DATA".RIO_06.FIRST_TANK.BWT_TEMP, 1 s
   "20_TANKS_IP_DATA_RIO_06_FIRST_TANK_DECK_IG_PRESS" : Real = PLC "20_TANKS_IP_DATA".RIO_06.FIRST_TANK.DECK_IG_PRESS, 1 s
   "20_TANKS_IP_DATA_RIO_06_FIRST_TANK_GTT_ISOL_VALVE_CLSD" : Bool = PLC "20_TANKS_IP_DATA".RIO_06.FIRST_TANK.GTT_ISOL_VALVE_CLSD, 1 s
   "20_TANKS_IP_DATA_RIO_06_FIRST_TANK_GTT_ISOL_VALVE_OPEN" : Bool = PLC "20_TANKS_IP_DATA".RIO_06.FIRST_TANK.GTT_ISOL_VALVE_OPEN, 1 s
   "20_TANKS_IP_DATA_RIO_06_FIRST_TANK_MBG_FLOW" : Real = PLC "20_TANKS_IP_DATA".RIO_06.FIRST_TANK.MBG_FLOW, 1 s
   "20_TANKS_IP_DATA_RIO_06_FIRST_TANK_O2_MONITOR" : Real = PLC "20_TANKS_IP_DATA".RIO_06.FIRST_TANK.O2_MONITOR, 1 s
   "20_TANKS_IP_DATA_RIO_06_FIRST_TANK_TANKS_PRESS" : Real = PLC "20_TANKS_IP_DATA".RIO_06.FIRST_TANK.TANKS_PRESS, 1 s
   "20_TANKS_IP_DATA_RIO_06_FIRST_TANK_USD_FLOW" : Real = PLC "20_TANKS_IP_DATA".RIO_06.FIRST_TANK.USD_FLOW, 1 s
   "20_TANKS_IP_DATA_RIO_06_SECOND_TANK_BWT_DO" : Real = PLC "20_TANKS_IP_DATA".RIO_06.SECOND_TANK.BWT_DO, 1 s
   "20_TANKS_IP_DATA_RIO_06_SECOND_TANK_BWT_LEVEL" : Real = PLC "20_TANKS_IP_DATA".RIO_06.SECOND_TANK.BWT_LEVEL, 1 s
   "20_TANKS_IP_DATA_RIO_06_SECOND_TANK_BWT_LEVEL_HIHI" : Bool = PLC "20_TANKS_IP_DATA".RIO_06.SECOND_TANK.BWT_LEVEL_HIHI, 1 s
   "20_TANKS_IP_DATA_RIO_06_SECOND_TANK_BWT_PH" : Real = PLC "20_TANKS_IP_DATA".RIO_06.SECOND_TANK.BWT_PH, 1 s
   "20_TANKS_IP_DATA_RIO_06_SECOND_TANK_BWT_TEMP" : Real = PLC "20_TANKS_IP_DATA".RIO_06.SECOND_TANK.BWT_TEMP, 1 s
   "20_TANKS_IP_DATA_RIO_06_SECOND_TANK_GTT_ISOL_VALVE_CLSD" : Bool = PLC "20_TANKS_IP_DATA".RIO_06.SECOND_TANK.GTT_ISOL_VALVE_CLSD, 1 s
   "20_TANKS_IP_DATA_RIO_06_SECOND_TANK_GTT_ISOL_VALVE_OPEN" : Bool = PLC "20_TANKS_IP_DATA".RIO_06.SECOND_TANK.GTT_ISOL_VALVE_OPEN, 1 s
   "20_TANKS_IP_DATA_RIO_06_SECOND_TANK_MBG_FLOW" : Real = PLC "20_TANKS_IP_DATA".RIO_06.SECOND_TANK.MBG_FLOW, 1 s
   "20_TANKS_IP_DATA_RIO_06_SECOND_TANK_TANKS_PRESS" : Real = PLC "20_TANKS_IP_DATA".RIO_06.SECOND_TANK.TANKS_PRESS, 1 s
   "20_TANKS_IP_DATA_RIO_06_SECOND_TANK_USD_FLOW" : Real = PLC "20_TANKS_IP_DATA".RIO_06.SECOND_TANK.USD_FLOW, 1 s
   "20_TANKS_IP_DATA_RIO_07_FIRST_TANK_BWT_DO" : Real = PLC "20_TANKS_IP_DATA".RIO_07.FIRST_TANK.BWT_DO, 1 s
   "20_TANKS_IP_DATA_RIO_07_FIRST_TANK_BWT_LEVEL" : Real = PLC "20_TANKS_IP_DATA".RIO_07.FIRST_TANK.BWT_LEVEL, 1 s
   "20_TANKS_IP_DATA_RIO_07_FIRST_TANK_BWT_LEVEL_HIHI" : Bool = PLC "20_TANKS_IP_DATA".RIO_07.FIRST_TANK.BWT_LEVEL_HIHI, 1 s
   "20_TANKS_IP_DATA_RIO_07_FIRST_TANK_BWT_PH" : Real = PLC "20_TANKS_IP_DATA".RIO_07.FIRST_TANK.BWT_PH, 1 s
   "20_TANKS_IP_DATA_RIO_07_FIRST_TANK_BWT_TEMP" : Real = PLC "20_TANKS_IP_DATA".RIO_07.FIRST_TANK.BWT_TEMP, 1 s
   "20_TANKS_IP_DATA_RIO_07_FIRST_TANK_DECK_IG_PRESS" : Real = PLC "20_TANKS_IP_DATA".RIO_07.FIRST_TANK.DECK_IG_PRESS, 1 s
   "20_TANKS_IP_DATA_RIO_07_FIRST_TANK_GTT_ISOL_VALVE_CLSD" : Bool = PLC "20_TANKS_IP_DATA".RIO_07.FIRST_TANK.GTT_ISOL_VALVE_CLSD, 1 s
   "20_TANKS_IP_DATA_RIO_07_FIRST_TANK_GTT_ISOL_VALVE_OPEN" : Bool = PLC "20_TANKS_IP_DATA".RIO_07.FIRST_TANK.GTT_ISOL_VALVE_OPEN, 1 s
   "20_TANKS_IP_DATA_RIO_07_FIRST_TANK_MBG_FLOW" : Real = PLC "20_TANKS_IP_DATA".RIO_07.FIRST_TANK.MBG_FLOW, 1 s
   "20_TANKS_IP_DATA_RIO_07_FIRST_TANK_O2_MONITOR" : Real = PLC "20_TANKS_IP_DATA".RIO_07.FIRST_TANK.O2_MONITOR, 1 s
   "20_TANKS_IP_DATA_RIO_07_FIRST_TANK_TANKS_PRESS" : Real = PLC "20_TANKS_IP_DATA".RIO_07.FIRST_TANK.TANKS_PRESS, 1 s
   "20_TANKS_IP_DATA_RIO_07_FIRST_TANK_USD_FLOW" : Real = PLC "20_TANKS_IP_DATA".RIO_07.FIRST_TANK.USD_FLOW, 1 s
   "2019_AUT_MAN_CNTRL_PORT_GTT_VLV_MAN" : Bool = PLC "2019_AUT_MAN_CNTRL".PORT_GTT_VLV_MAN AT %DB1.DBW0, 1 s
   "2019_AUT_MAN_CNTRL_STBD_GTT_VLV_MAN" : Bool = PLC "2019_AUT_MAN_CNTRL".STBD_GTT_VLV_MAN AT %DB1.DBW0, 1 s
   "2060_Alarm_Data_BTCS_ALARM_WORD_1" : Word = PLC "2060_Alarm_Data".BTCS_ALARM_WORD_01 AT %DB2060.DBW0, 1 s
   "2060_Alarm_Data_BTCS_ALARM_WORD_2" : Word = PLC "2060_Alarm_Data".BTCS_ALARM_WORD_02 AT %DB2060.DBW2, 1 s
   "2060_Alarm_Data_BTCS_ALARM_WORD_3" : Word = PLC "2060_Alarm_Data".BTCS_ALARM_WORD_03 AT %DB2060.DBW4, 1 s
   "2060_Alarm_Data_BTCS_ALARM_WORD_4" : Word = PLC "2060_Alarm_Data".BTCS_ALARM_WORD_04 AT %DB2060.DBW6, 1 s
   "2060_Alarm_Data_BTCS_ALARM_WORD_5" : Word = PLC "2060_Alarm_Data".BTCS_ALARM_WORD_05 AT %DB2060.DBW8, 1 s
   "2060_Alarm_Data_BTCS_ALARM_WORD_6" : Word = PLC "2060_Alarm_Data".BTCS_ALARM_WORD_06 AT %DB2060.DBW10, 1 s
   "2060_Alarm_Data_BTCS_ALARM_WORD_7" : Word = PLC "2060_Alarm_Data".BTCS_ALARM_WORD_07 AT %DB2060.DBW12, 1 s
   "2060_Alarm_Data_BTCS_ALARM_WORD_8" : Word = PLC "2060_Alarm_Data".BTCS_ALARM_WORD_08 AT %DB2060.DBW14, 1 s
   "2062_Warning_Data_Alarm Tank APT" : Bool = PLC "2062_Warning_Data"."Alarm Tank APT" AT %DB2062.DBX23.6, 1 s
   "2062_Warning_Data_Alarm Tank FPT" : Bool = PLC "2062_Warning_Data"."Alarm Tank FPT" AT %DB2062.DBX22.1, 1 s
   "2062_Warning_Data_Alarm Tank P1" : Bool = PLC "2062_Warning_Data"."Alarm Tank P1" AT %DB2062.DBX22.2, 1 s
   "2062_Warning_Data_Alarm Tank P2" : Bool = PLC "2062_Warning_Data"."Alarm Tank P2" AT %DB2062.DBX22.4, 1 s
   "2062_Warning_Data_Alarm Tank P3" : Bool = PLC "2062_Warning_Data"."Alarm Tank P3" AT %DB2062.DBX22.6, 1 s
   "2062_Warning_Data_Alarm Tank P4" : Bool = PLC "2062_Warning_Data"."Alarm Tank P4" AT %DB2062.DBX23.0, 1 s
   "2062_Warning_Data_Alarm Tank P5" : Bool = PLC "2062_Warning_Data"."Alarm Tank P5" AT %DB2062.DBX23.2, 1 s
   "2062_Warning_Data_Alarm Tank P6" : Bool = PLC "2062_Warning_Data"."Alarm Tank P6" AT %DB2062.DBX23.4, 1 s
   "2062_Warning_Data_Alarm Tank S1" : Bool = PLC "2062_Warning_Data"."Alarm Tank S1" AT %DB2062.DBX22.3, 1 s
   "2062_Warning_Data_Alarm Tank S2" : Bool = PLC "2062_Warning_Data"."Alarm Tank S2" AT %DB2062.DBX22.5, 1 s
   "2062_Warning_Data_Alarm Tank S3" : Bool = PLC "2062_Warning_Data"."Alarm Tank S3" AT %DB2062.DBX22.7, 1 s
   "2062_Warning_Data_Alarm Tank S4" : Bool = PLC "2062_Warning_Data"."Alarm Tank S4" AT %DB2062.DBX23.1, 1 s
   "2062_Warning_Data_Alarm Tank S5" : Bool = PLC "2062_Warning_Data"."Alarm Tank S5" AT %DB2062.DBX23.3, 1 s
   "2062_Warning_Data_Alarm Tank S6" : Bool = PLC "2062_Warning_Data"."Alarm Tank S6" AT %DB2062.DBX23.5, 1 s
   "2062_Warning_Data_BTCS_WARNING_WORD_09" : Word = PLC "2062_Warning_Data".BTCS_WARNING_WORD_09 AT %DB2062.DBW16, 1 s
   "2062_Warning_Data_BTCS_WARNING_WORD_1" : Word = PLC "2062_Warning_Data".BTCS_WARNING_WORD_01 AT %DB2062.DBW0, 1 s
   "2062_Warning_Data_BTCS_WARNING_WORD_10" : Word = PLC "2062_Warning_Data".BTCS_WARNING_WORD_10 AT %DB2062.DBW18, 1 s
   "2062_Warning_Data_BTCS_WARNING_WORD_11" : Word = PLC "2062_Warning_Data".BTCS_WARNING_WORD_11 AT %DB2062.DBW20, 1 s
   "2062_Warning_Data_BTCS_WARNING_WORD_12" : Word = PLC "2062_Warning_Data".BTCS_WARNING_WORD_12 AT %DB2062.DBW362, 1 s